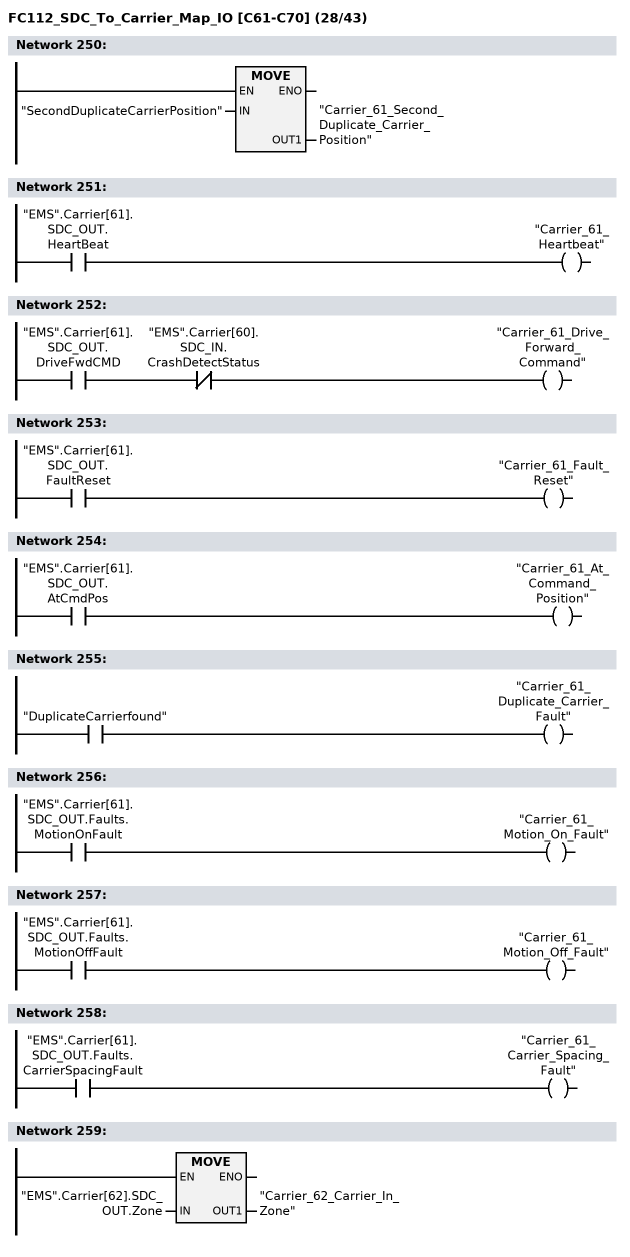
   RUNG wire#powerrail
      Move(in := "SecondDuplicateCarrierPosition", out1 => "Carrier_61_Second_Duplicate_Carrier_Position")
   END_RUNG
   // the same network as SCL:
   "Carrier_61_Second_Duplicate_Carrier_Position" := "SecondDuplicateCarrierPosition";
END_REGION

REGION Network 251
   RUNG wire#powerrail
      Contact( "EMS".Carrier[61].SDC_OUT.HeartBeat )
      Coil( "Carrier_61_Heartbeat" )
   END_RUNG
   // the same network as SCL:
   "Carrier_61_Heartbeat" := "EMS".Carrier[61].SDC_OUT.HeartBeat;
END_REGION

REGION Network 252
   RUNG wire#powerrail
      Contact( "EMS".Carrier[61].SDC_OUT.DriveFwdCMD )
      I_Contact( "EMS".Carrier[60].SDC_IN.CrashDetectStatus )
      Coil( "Carrier_61_Drive_Forward_Command" )
   END_RUNG
   // the same network as SCL:
   "Carrier_61_Drive_Forward_Command" := "EMS".Carrier[61].SDC_OUT.DriveFwdCMD AND NOT "EMS".Carrier[60].SDC_IN.CrashDetectStatus;
END_REGION

REGION Network 253
   RUNG wire#powerrail
      Contact( "EMS".Carrier[61].SDC_OUT.FaultReset )
      Coil( "Carrier_61_Fault_Reset" )
   END_RUNG
   // the same network as SCL:
   "Carrier_61_Fault_Reset" := "EMS".Carrier[61].SDC_OUT.FaultReset;
END_REGION

REGION Network 254
   RUNG wire#powerrail
      Contact( "EMS".Carrier[61].SDC_OUT.AtCmdPos )
      Coil( "Carrier_61_At_Command_Position" )
   END_RUNG
   // the same network as SCL:
   "Carrier_61_At_Command_Position" := "EMS".Carrier[61].SDC_OUT.AtCmdPos;
END_REGION

REGION Network 255
   RUNG wire#powerrail
      Contact( "DuplicateCarrierfound" )
      Coil( "Carrier_61_Duplicate_Carrier_Fault" )
   END_RUNG
   // the same network as SCL:
   "Carrier_61_Duplicate_Carrier_Fault" := "DuplicateCarrierfound";
END_REGION

REGION Network 256
   RUNG wire#powerrail
      Contact( "EMS".Carrier[61].SDC_OUT.Faults.MotionOnFault )
      Coil( "Carrier_61_Motion_On_Fault" )
   END_RUNG
   // the same network as SCL:
   "Carrier_61_Motion_On_Fault" := "EMS".Carrier[61].SDC_OUT.Faults.MotionOnFault;
END_REGION

REGION Network 257
   RUNG wire#powerrail
      Contact( "EMS".Carrier[61].SDC_OUT.Faults.MotionOffFault )
      Coil( "Carrier_61_Motion_Off_Fault" )
   END_RUNG
   // the same network as SCL:
   "Carrier_61_Motion_Off_Fault" := "EMS".Carrier[61].SDC_OUT.Faults.MotionOffFault;
END_REGION

REGION Network 258
   RUNG wire#powerrail
      Contact( "EMS".Carrier[61].SDC_OUT.Faults.CarrierSpacingFault )
      Coil( "Carrier_61_Carrier_Spacing_Fault" )
   END_RUNG
   // the same network as SCL:
   "Carrier_61_Carrier_Spacing_Fault" := "EMS".Carrier[61].SDC_OUT.Faults.CarrierSpacingFault;
END_REGION

REGION Network 259
   RUNG wire#powerrail
      Move(in := "EMS".Carrier[62].SDC_OUT.Zone, out1 => "Carrier_62_Carrier_In_Zone")
   END_RUNG
   // the same network as SCL:
   "Carrier_62_Carrier_In_Zone" := "EMS".Carrier[62].SDC_OUT.Zone;
END_REGION

REGION Network 260
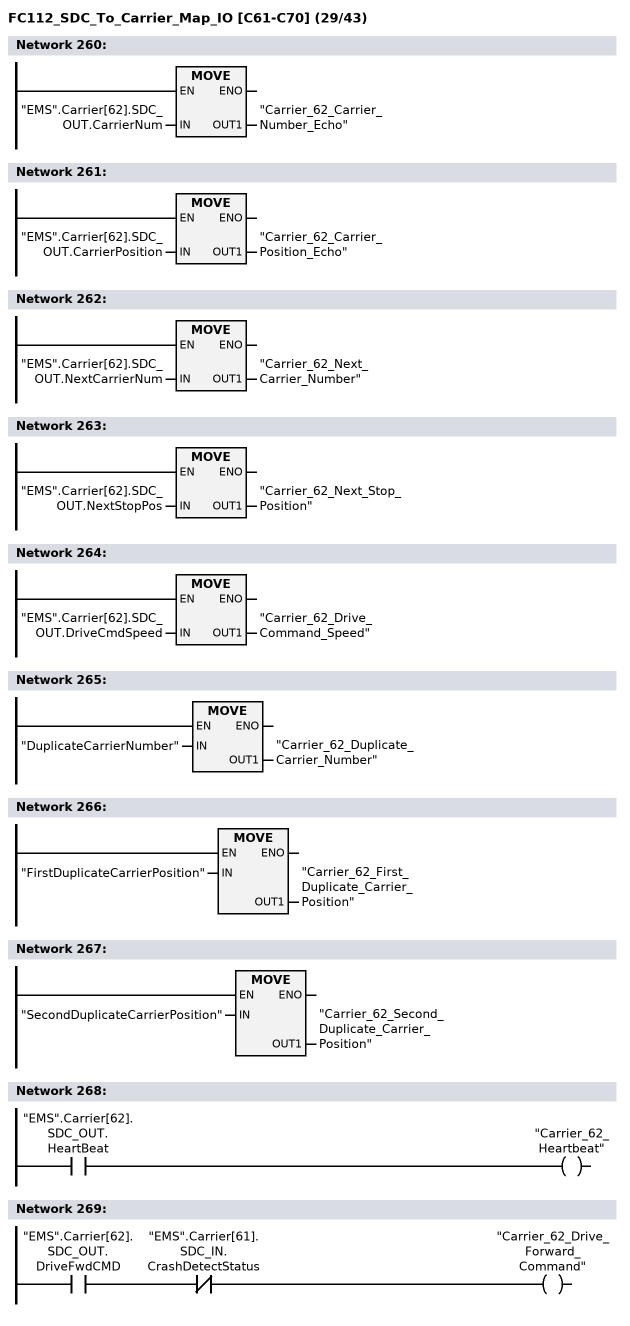
   RUNG wire#powerrail
      Move(in := "EMS".Carrier[62].SDC_OUT.CarrierNum, out1 => "Carrier_62_Carrier_Number_Echo")
   END_RUNG
   // the same network as SCL:
   "Carrier_62_Carrier_Number_Echo" := "EMS".Carrier[62].SDC_OUT.CarrierNum;
END_REGION

REGION Network 261
   RUNG wire#powerrail
      Move(in := "EMS".Carrier[62].SDC_OUT.CarrierPosition, out1 => "Carrier_62_Carrier_Position_Echo")
   END_RUNG
   // the same network as SCL:
   "Carrier_62_Carrier_Position_Echo" := "EMS".Carrier[62].SDC_OUT.CarrierPosition;
END_REGION

REGION Network 262
   RUNG wire#powerrail
      Move(in := "EMS".Carrier[62].SDC_OUT.NextCarrierNum, out1 => "Carrier_62_Next_Carrier_Number")
   END_RUNG
   // the same network as SCL:
   "Carrier_62_Next_Carrier_Number" := "EMS".Carrier[62].SDC_OUT.NextCarrierNum;
END_REGION

REGION Network 263
   RUNG wire#powerrail
      Move(in := "EMS".Carrier[62].SDC_OUT.NextStopPos, out1 => "Carrier_62_Next_Stop_Position")
   END_RUNG
   // the same network as SCL:
   "Carrier_62_Next_Stop_Position" := "EMS".Carrier[62].SDC_OUT.NextStopPos;
END_REGION

REGION Network 264
   RUNG wire#powerrail
      Move(in := "EMS".Carrier[62].SDC_OUT.DriveCmdSpeed, out1 => "Carrier_62_Drive_Command_Speed")
   END_RUNG
   // the same network as SCL:
   "Carrier_62_Drive_Command_Speed" := "EMS".Carrier[62].SDC_OUT.DriveCmdSpeed;
END_REGION

REGION Network 265
   RUNG wire#powerrail
      Move(in := "DuplicateCarrierNumber", out1 => "Carrier_62_Duplicate_Carrier_Number")
   END_RUNG
   // the same network as SCL:
   "Carrier_62_Duplicate_Carrier_Number" := "DuplicateCarrierNumber";
END_REGION

REGION Network 266
   RUNG wire#powerrail
      Move(in := "FirstDuplicateCarrierPosition", out1 => "Carrier_62_First_Duplicate_Carrier_Position")
   END_RUNG
   // the same network as SCL:
   "Carrier_62_First_Duplicate_Carrier_Position" := "FirstDuplicateCarrierPosition";
END_REGION

REGION Network 267
   RUNG wire#powerrail
      Move(in := "SecondDuplicateCarrierPosition", out1 => "Carrier_62_Second_Duplicate_Carrier_Position")
   END_RUNG
   // the same network as SCL:
   "Carrier_62_Second_Duplicate_Carrier_Position" := "SecondDuplicateCarrierPosition";
END_REGION

REGION Network 268
   RUNG wire#powerrail
      Contact( "EMS".Carrier[62].SDC_OUT.HeartBeat )
      Coil( "Carrier_62_Heartbeat" )
   END_RUNG
   // the same network as SCL:
   "Carrier_62_Heartbeat" := "EMS".Carrier[62].SDC_OUT.HeartBeat;
END_REGION

REGION Network 269
   RUNG wire#powerrail
      Contact( "EMS".Carrier[62].SDC_OUT.DriveFwdCMD )
      I_Contact( "EMS".Carrier[61].SDC_IN.CrashDetectStatus )
      Coil( "Carrier_62_Drive_Forward_Command" )
   END_RUNG
   // the same network as SCL:
   "Carrier_62_Drive_Forward_Command" := "EMS".Carrier[62].SDC_OUT.DriveFwdCMD AND NOT "EMS".Carrier[61].SDC_IN.CrashDetectStatus;
END_REGION

REGION Network 270
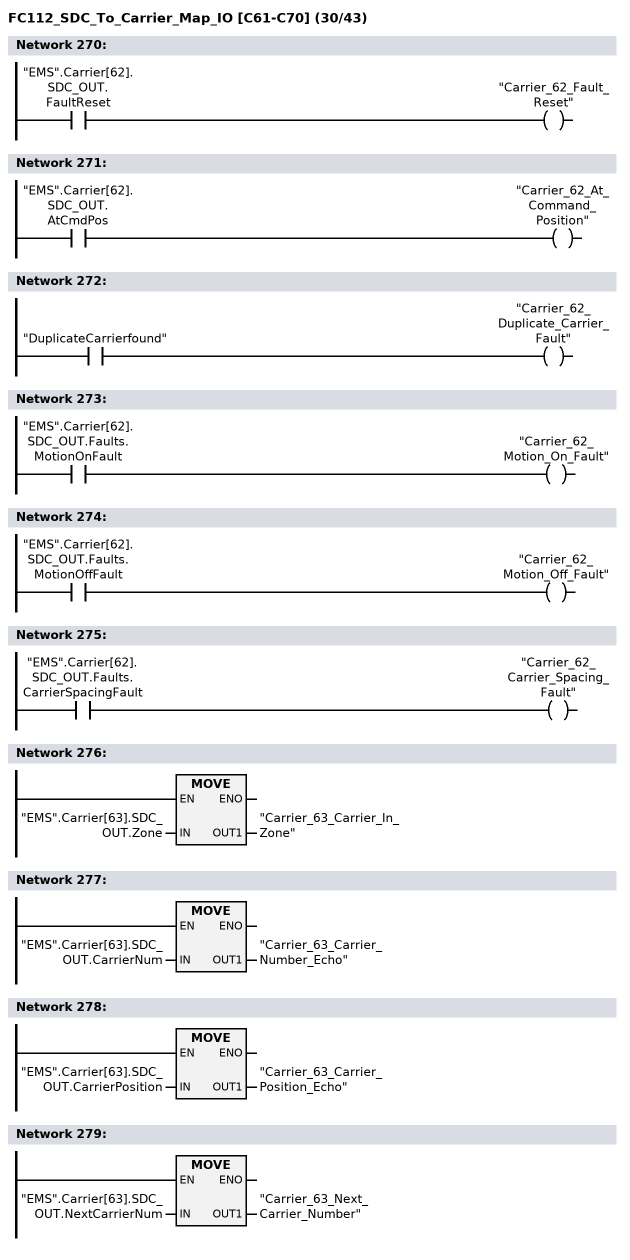
   RUNG wire#powerrail
      Contact( "EMS".Carrier[62].SDC_OUT.FaultReset )
      Coil( "Carrier_62_Fault_Reset" )
   END_RUNG
   // the same network as SCL:
   "Carrier_62_Fault_Reset" := "EMS".Carrier[62].SDC_OUT.FaultReset;
END_REGION

REGION Network 271
   RUNG wire#powerrail
      Contact( "EMS".Carrier[62].SDC_OUT.AtCmdPos )
      Coil( "Carrier_62_At_Command_Position" )
   END_RUNG
   // the same network as SCL:
   "Carrier_62_At_Command_Position" := "EMS".Carrier[62].SDC_OUT.AtCmdPos;
END_REGION

REGION Network 272
   RUNG wire#powerrail
      Contact( "DuplicateCarrierfound" )
      Coil( "Carrier_62_Duplicate_Carrier_Fault" )
   END_RUNG
   // the same network as SCL:
   "Carrier_62_Duplicate_Carrier_Fault" := "DuplicateCarrierfound";
END_REGION

REGION Network 273
   RUNG wire#powerrail
      Contact( "EMS".Carrier[62].SDC_OUT.Faults.MotionOnFault )
      Coil( "Carrier_62_Motion_On_Fault" )
   END_RUNG
   // the same network as SCL:
   "Carrier_62_Motion_On_Fault" := "EMS".Carrier[62].SDC_OUT.Faults.MotionOnFault;
END_REGION

REGION Network 274
   RUNG wire#powerrail
      Contact( "EMS".Carrier[62].SDC_OUT.Faults.MotionOffFault )
      Coil( "Carrier_62_Motion_Off_Fault" )
   END_RUNG
   // the same network as SCL:
   "Carrier_62_Motion_Off_Fault" := "EMS".Carrier[62].SDC_OUT.Faults.MotionOffFault;
END_REGION

REGION Network 275
   RUNG wire#powerrail
      Contact( "EMS".Carrier[62].SDC_OUT.Faults.CarrierSpacingFault )
      Coil( "Carrier_62_Carrier_Spacing_Fault" )
   END_RUNG
   // the same network as SCL:
   "Carrier_62_Carrier_Spacing_Fault" := "EMS".Carrier[62].SDC_OUT.Faults.CarrierSpacingFault;
END_REGION

REGION Network 276
   RUNG wire#powerrail
      Move(in := "EMS".Carrier[63].SDC_OUT.Zone, out1 => "Carrier_63_Carrier_In_Zone")
   END_RUNG
   // the same network as SCL:
   "Carrier_63_Carrier_In_Zone" := "EMS".Carrier[63].SDC_OUT.Zone;
END_REGION

REGION Network 277
   RUNG wire#powerrail
      Move(in := "EMS".Carrier[63].SDC_OUT.CarrierNum, out1 => "Carrier_63_Carrier_Number_Echo")
   END_RUNG
   // the same network as SCL:
   "Carrier_63_Carrier_Number_Echo" := "EMS".Carrier[63].SDC_OUT.CarrierNum;
END_REGION

REGION Network 278
   RUNG wire#powerrail
      Move(in := "EMS".Carrier[63].SDC_OUT.CarrierPosition, out1 => "Carrier_63_Carrier_Position_Echo")
   END_RUNG
   // the same network as SCL:
   "Carrier_63_Carrier_Position_Echo" := "EMS".Carrier[63].SDC_OUT.CarrierPosition;
END_REGION

REGION Network 279
   RUNG wire#powerrail
      Move(in := "EMS".Carrier[63].SDC_OUT.NextCarrierNum, out1 => "Carrier_63_Next_Carrier_Number")
   END_RUNG
   // the same network as SCL:
   "Carrier_63_Next_Carrier_Number" := "EMS".Carrier[63].SDC_OUT.NextCarrierNum;
END_REGION

REGION Network 280
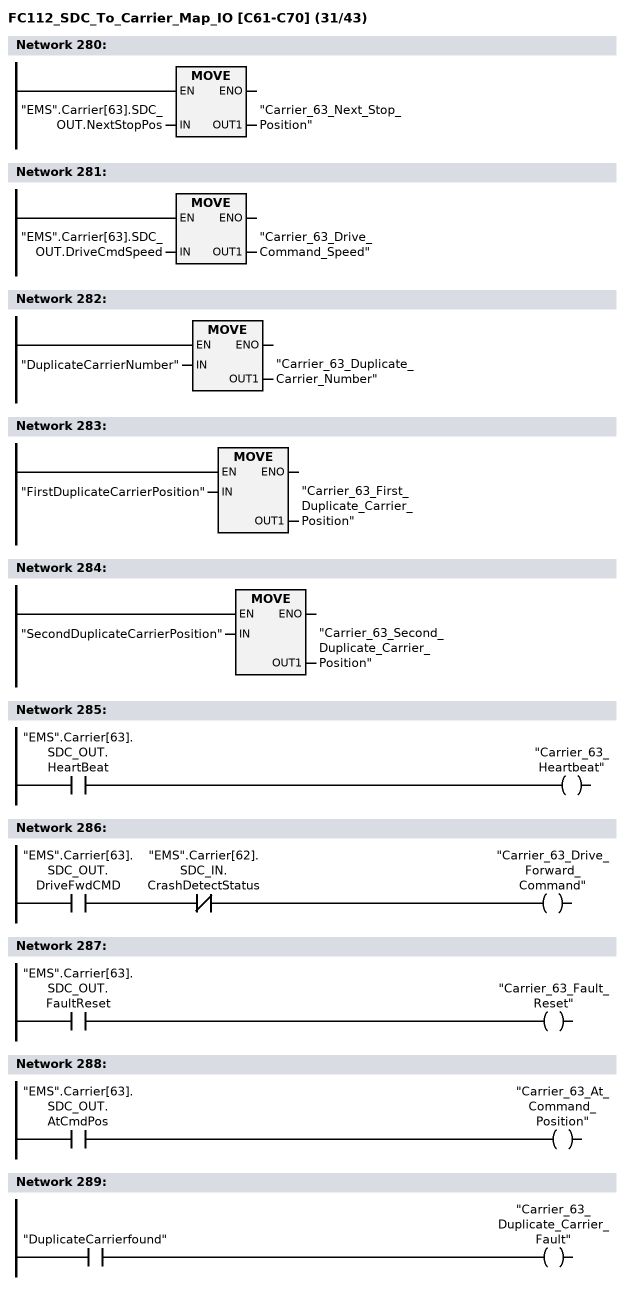
   RUNG wire#powerrail
      Move(in := "EMS".Carrier[63].SDC_OUT.NextStopPos, out1 => "Carrier_63_Next_Stop_Position")
   END_RUNG
   // the same network as SCL:
   "Carrier_63_Next_Stop_Position" := "EMS".Carrier[63].SDC_OUT.NextStopPos;
END_REGION

REGION Network 281
   RUNG wire#powerrail
      Move(in := "EMS".Carrier[63].SDC_OUT.DriveCmdSpeed, out1 => "Carrier_63_Drive_Command_Speed")
   END_RUNG
   // the same network as SCL:
   "Carrier_63_Drive_Command_Speed" := "EMS".Carrier[63].SDC_OUT.DriveCmdSpeed;
END_REGION

REGION Network 282
   RUNG wire#powerrail
      Move(in := "DuplicateCarrierNumber", out1 => "Carrier_63_Duplicate_Carrier_Number")
   END_RUNG
   // the same network as SCL:
   "Carrier_63_Duplicate_Carrier_Number" := "DuplicateCarrierNumber";
END_REGION

REGION Network 283
   RUNG wire#powerrail
      Move(in := "FirstDuplicateCarrierPosition", out1 => "Carrier_63_First_Duplicate_Carrier_Position")
   END_RUNG
   // the same network as SCL:
   "Carrier_63_First_Duplicate_Carrier_Position" := "FirstDuplicateCarrierPosition";
END_REGION

REGION Network 284
   RUNG wire#powerrail
      Move(in := "SecondDuplicateCarrierPosition", out1 => "Carrier_63_Second_Duplicate_Carrier_Position")
   END_RUNG
   // the same network as SCL:
   "Carrier_63_Second_Duplicate_Carrier_Position" := "SecondDuplicateCarrierPosition";
END_REGION

REGION Network 285
   RUNG wire#powerrail
      Contact( "EMS".Carrier[63].SDC_OUT.HeartBeat )
      Coil( "Carrier_63_Heartbeat" )
   END_RUNG
   // the same network as SCL:
   "Carrier_63_Heartbeat" := "EMS".Carrier[63].SDC_OUT.HeartBeat;
END_REGION

REGION Network 286
   RUNG wire#powerrail
      Contact( "EMS".Carrier[63].SDC_OUT.DriveFwdCMD )
      I_Contact( "EMS".Carrier[62].SDC_IN.CrashDetectStatus )
      Coil( "Carrier_63_Drive_Forward_Command" )
   END_RUNG
   // the same network as SCL:
   "Carrier_63_Drive_Forward_Command" := "EMS".Carrier[63].SDC_OUT.DriveFwdCMD AND NOT "EMS".Carrier[62].SDC_IN.CrashDetectStatus;
END_REGION

REGION Network 287
   RUNG wire#powerrail
      Contact( "EMS".Carrier[63].SDC_OUT.FaultReset )
      Coil( "Carrier_63_Fault_Reset" )
   END_RUNG
   // the same network as SCL:
   "Carrier_63_Fault_Reset" := "EMS".Carrier[63].SDC_OUT.FaultReset;
END_REGION

REGION Network 288
   RUNG wire#powerrail
      Contact( "EMS".Carrier[63].SDC_OUT.AtCmdPos )
      Coil( "Carrier_63_At_Command_Position" )
   END_RUNG
   // the same network as SCL:
   "Carrier_63_At_Command_Position" := "EMS".Carrier[63].SDC_OUT.AtCmdPos;
END_REGION

REGION Network 289
   RUNG wire#powerrail
      Contact( "DuplicateCarrierfound" )
      Coil( "Carrier_63_Duplicate_Carrier_Fault" )
   END_RUNG
   // the same network as SCL:
   "Carrier_63_Duplicate_Carrier_Fault" := "DuplicateCarrierfound";
END_REGION

REGION Network 290
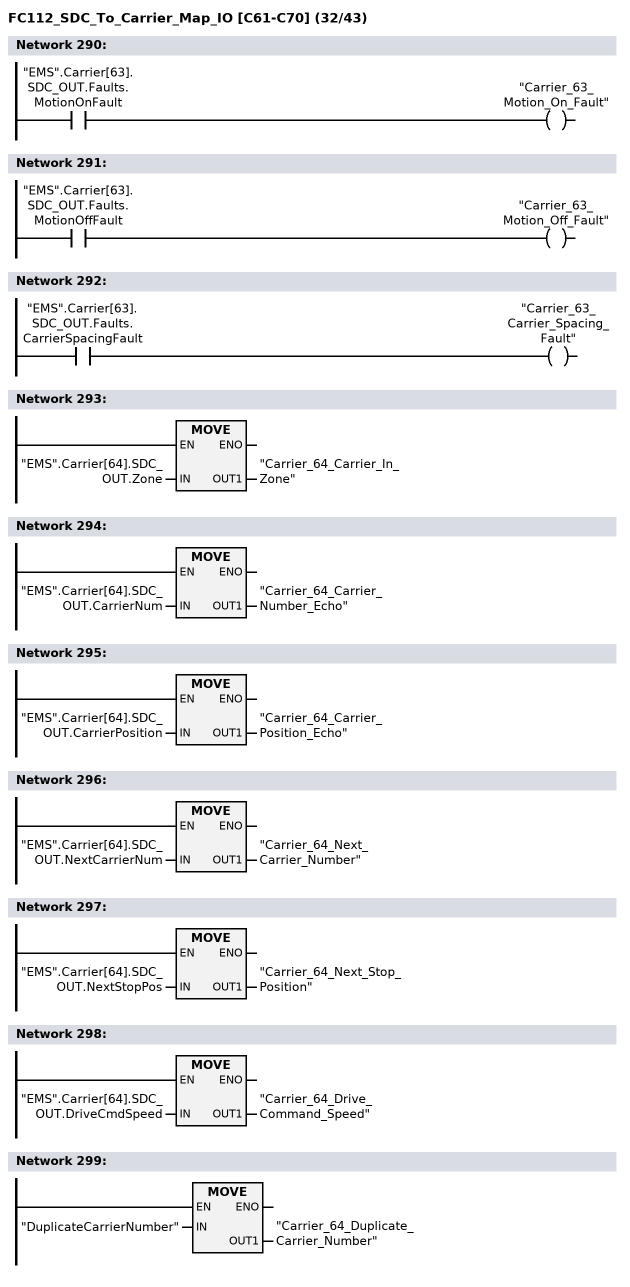
   RUNG wire#powerrail
      Contact( "EMS".Carrier[63].SDC_OUT.Faults.MotionOnFault )
      Coil( "Carrier_63_Motion_On_Fault" )
   END_RUNG
   // the same network as SCL:
   "Carrier_63_Motion_On_Fault" := "EMS".Carrier[63].SDC_OUT.Faults.MotionOnFault;
END_REGION

REGION Network 291
   RUNG wire#powerrail
      Contact( "EMS".Carrier[63].SDC_OUT.Faults.MotionOffFault )
      Coil( "Carrier_63_Motion_Off_Fault" )
   END_RUNG
   // the same network as SCL:
   "Carrier_63_Motion_Off_Fault" := "EMS".Carrier[63].SDC_OUT.Faults.MotionOffFault;
END_REGION

REGION Network 292
   RUNG wire#powerrail
      Contact( "EMS".Carrier[63].SDC_OUT.Faults.CarrierSpacingFault )
      Coil( "Carrier_63_Carrier_Spacing_Fault" )
   END_RUNG
   // the same network as SCL:
   "Carrier_63_Carrier_Spacing_Fault" := "EMS".Carrier[63].SDC_OUT.Faults.CarrierSpacingFault;
END_REGION

REGION Network 293
   RUNG wire#powerrail
      Move(in := "EMS".Carrier[64].SDC_OUT.Zone, out1 => "Carrier_64_Carrier_In_Zone")
   END_RUNG
   // the same network as SCL:
   "Carrier_64_Carrier_In_Zone" := "EMS".Carrier[64].SDC_OUT.Zone;
END_REGION

REGION Network 294
   RUNG wire#powerrail
      Move(in := "EMS".Carrier[64].SDC_OUT.CarrierNum, out1 => "Carrier_64_Carrier_Number_Echo")
   END_RUNG
   // the same network as SCL:
   "Carrier_64_Carrier_Number_Echo" := "EMS".Carrier[64].SDC_OUT.CarrierNum;
END_REGION

REGION Network 295
   RUNG wire#powerrail
      Move(in := "EMS".Carrier[64].SDC_OUT.CarrierPosition, out1 => "Carrier_64_Carrier_Position_Echo")
   END_RUNG
   // the same network as SCL:
   "Carrier_64_Carrier_Position_Echo" := "EMS".Carrier[64].SDC_OUT.CarrierPosition;
END_REGION

REGION Network 296
   RUNG wire#powerrail
      Move(in := "EMS".Carrier[64].SDC_OUT.NextCarrierNum, out1 => "Carrier_64_Next_Carrier_Number")
   END_RUNG
   // the same network as SCL:
   "Carrier_64_Next_Carrier_Number" := "EMS".Carrier[64].SDC_OUT.NextCarrierNum;
END_REGION

REGION Network 297
   RUNG wire#powerrail
      Move(in := "EMS".Carrier[64].SDC_OUT.NextStopPos, out1 => "Carrier_64_Next_Stop_Position")
   END_RUNG
   // the same network as SCL:
   "Carrier_64_Next_Stop_Position" := "EMS".Carrier[64].SDC_OUT.NextStopPos;
END_REGION

REGION Network 298
   RUNG wire#powerrail
      Move(in := "EMS".Carrier[64].SDC_OUT.DriveCmdSpeed, out1 => "Carrier_64_Drive_Command_Speed")
   END_RUNG
   // the same network as SCL:
   "Carrier_64_Drive_Command_Speed" := "EMS".Carrier[64].SDC_OUT.DriveCmdSpeed;
END_REGION

REGION Network 299
   RUNG wire#powerrail
      Move(in := "DuplicateCarrierNumber", out1 => "Carrier_64_Duplicate_Carrier_Number")
   END_RUNG
   // the same network as SCL:
   "Carrier_64_Duplicate_Carrier_Number" := "DuplicateCarrierNumber";
END_REGION

REGION Network 300
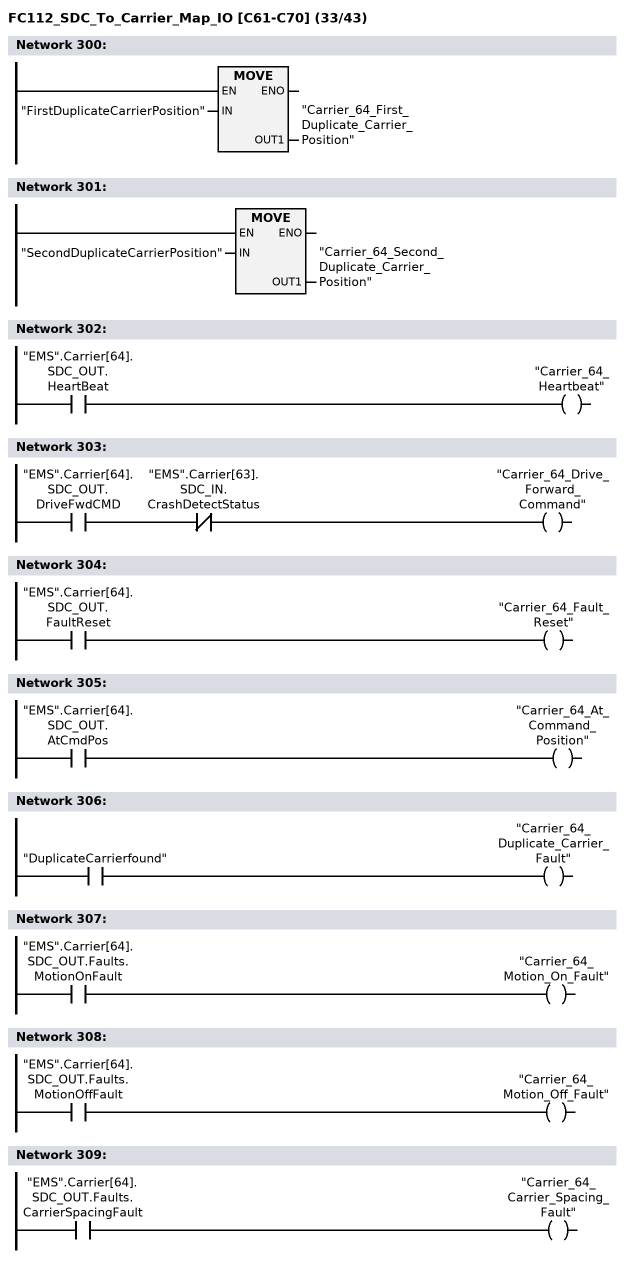
   RUNG wire#powerrail
      Move(in := "FirstDuplicateCarrierPosition", out1 => "Carrier_64_First_Duplicate_Carrier_Position")
   END_RUNG
   // the same network as SCL:
   "Carrier_64_First_Duplicate_Carrier_Position" := "FirstDuplicateCarrierPosition";
END_REGION

REGION Network 301
   RUNG wire#powerrail
      Move(in := "SecondDuplicateCarrierPosition", out1 => "Carrier_64_Second_Duplicate_Carrier_Position")
   END_RUNG
   // the same network as SCL:
   "Carrier_64_Second_Duplicate_Carrier_Position" := "SecondDuplicateCarrierPosition";
END_REGION

REGION Network 302
   RUNG wire#powerrail
      Contact( "EMS".Carrier[64].SDC_OUT.HeartBeat )
      Coil( "Carrier_64_Heartbeat" )
   END_RUNG
   // the same network as SCL:
   "Carrier_64_Heartbeat" := "EMS".Carrier[64].SDC_OUT.HeartBeat;
END_REGION

REGION Network 303
   RUNG wire#powerrail
      Contact( "EMS".Carrier[64].SDC_OUT.DriveFwdCMD )
      I_Contact( "EMS".Carrier[63].SDC_IN.CrashDetectStatus )
      Coil( "Carrier_64_Drive_Forward_Command" )
   END_RUNG
   // the same network as SCL:
   "Carrier_64_Drive_Forward_Command" := "EMS".Carrier[64].SDC_OUT.DriveFwdCMD AND NOT "EMS".Carrier[63].SDC_IN.CrashDetectStatus;
END_REGION

REGION Network 304
   RUNG wire#powerrail
      Contact( "EMS".Carrier[64].SDC_OUT.FaultReset )
      Coil( "Carrier_64_Fault_Reset" )
   END_RUNG
   // the same network as SCL:
   "Carrier_64_Fault_Reset" := "EMS".Carrier[64].SDC_OUT.FaultReset;
END_REGION

REGION Network 305
   RUNG wire#powerrail
      Contact( "EMS".Carrier[64].SDC_OUT.AtCmdPos )
      Coil( "Carrier_64_At_Command_Position" )
   END_RUNG
   // the same network as SCL:
   "Carrier_64_At_Command_Position" := "EMS".Carrier[64].SDC_OUT.AtCmdPos;
END_REGION

REGION Network 306
   RUNG wire#powerrail
      Contact( "DuplicateCarrierfound" )
      Coil( "Carrier_64_Duplicate_Carrier_Fault" )
   END_RUNG
   // the same network as SCL:
   "Carrier_64_Duplicate_Carrier_Fault" := "DuplicateCarrierfound";
END_REGION

REGION Network 307
   RUNG wire#powerrail
      Contact( "EMS".Carrier[64].SDC_OUT.Faults.MotionOnFault )
      Coil( "Carrier_64_Motion_On_Fault" )
   END_RUNG
   // the same network as SCL:
   "Carrier_64_Motion_On_Fault" := "EMS".Carrier[64].SDC_OUT.Faults.MotionOnFault;
END_REGION

REGION Network 308
   RUNG wire#powerrail
      Contact( "EMS".Carrier[64].SDC_OUT.Faults.MotionOffFault )
      Coil( "Carrier_64_Motion_Off_Fault" )
   END_RUNG
   // the same network as SCL:
   "Carrier_64_Motion_Off_Fault" := "EMS".Carrier[64].SDC_OUT.Faults.MotionOffFault;
END_REGION

REGION Network 309
   RUNG wire#powerrail
      Contact( "EMS".Carrier[64].SDC_OUT.Faults.CarrierSpacingFault )
      Coil( "Carrier_64_Carrier_Spacing_Fault" )
   END_RUNG
   // the same network as SCL:
   "Carrier_64_Carrier_Spacing_Fault" := "EMS".Carrier[64].SDC_OUT.Faults.CarrierSpacingFault;
END_REGION

REGION Network 310
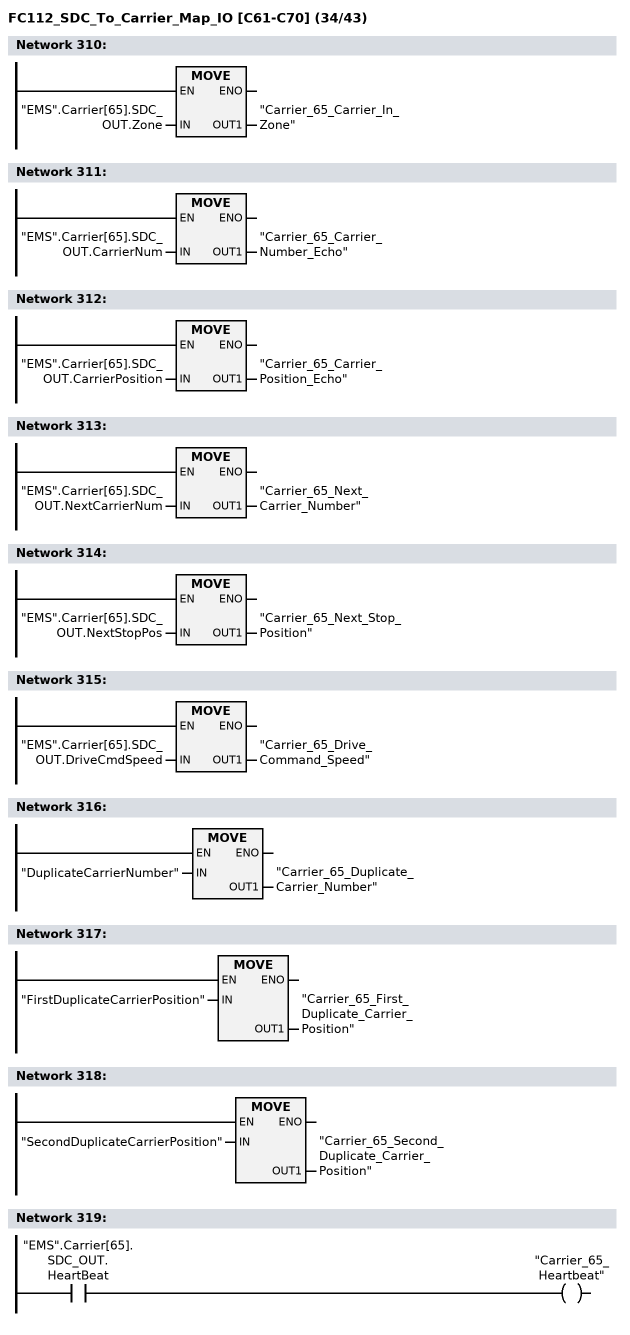
   RUNG wire#powerrail
      Move(in := "EMS".Carrier[65].SDC_OUT.Zone, out1 => "Carrier_65_Carrier_In_Zone")
   END_RUNG
   // the same network as SCL:
   "Carrier_65_Carrier_In_Zone" := "EMS".Carrier[65].SDC_OUT.Zone;
END_REGION

REGION Network 311
   RUNG wire#powerrail
      Move(in := "EMS".Carrier[65].SDC_OUT.CarrierNum, out1 => "Carrier_65_Carrier_Number_Echo")
   END_RUNG
   // the same network as SCL:
   "Carrier_65_Carrier_Number_Echo" := "EMS".Carrier[65].SDC_OUT.CarrierNum;
END_REGION

REGION Network 312
   RUNG wire#powerrail
      Move(in := "EMS".Carrier[65].SDC_OUT.CarrierPosition, out1 => "Carrier_65_Carrier_Position_Echo")
   END_RUNG
   // the same network as SCL:
   "Carrier_65_Carrier_Position_Echo" := "EMS".Carrier[65].SDC_OUT.CarrierPosition;
END_REGION

REGION Network 313
   RUNG wire#powerrail
      Move(in := "EMS".Carrier[65].SDC_OUT.NextCarrierNum, out1 => "Carrier_65_Next_Carrier_Number")
   END_RUNG
   // the same network as SCL:
   "Carrier_65_Next_Carrier_Number" := "EMS".Carrier[65].SDC_OUT.NextCarrierNum;
END_REGION

REGION Network 314
   RUNG wire#powerrail
      Move(in := "EMS".Carrier[65].SDC_OUT.NextStopPos, out1 => "Carrier_65_Next_Stop_Position")
   END_RUNG
   // the same network as SCL:
   "Carrier_65_Next_Stop_Position" := "EMS".Carrier[65].SDC_OUT.NextStopPos;
END_REGION

REGION Network 315
   RUNG wire#powerrail
      Move(in := "EMS".Carrier[65].SDC_OUT.DriveCmdSpeed, out1 => "Carrier_65_Drive_Command_Speed")
   END_RUNG
   // the same network as SCL:
   "Carrier_65_Drive_Command_Speed" := "EMS".Carrier[65].SDC_OUT.DriveCmdSpeed;
END_REGION

REGION Network 316
   RUNG wire#powerrail
      Move(in := "DuplicateCarrierNumber", out1 => "Carrier_65_Duplicate_Carrier_Number")
   END_RUNG
   // the same network as SCL:
   "Carrier_65_Duplicate_Carrier_Number" := "DuplicateCarrierNumber";
END_REGION

REGION Network 317
   RUNG wire#powerrail
      Move(in := "FirstDuplicateCarrierPosition", out1 => "Carrier_65_First_Duplicate_Carrier_Position")
   END_RUNG
   // the same network as SCL:
   "Carrier_65_First_Duplicate_Carrier_Position" := "FirstDuplicateCarrierPosition";
END_REGION

REGION Network 318
   RUNG wire#powerrail
      Move(in := "SecondDuplicateCarrierPosition", out1 => "Carrier_65_Second_Duplicate_Carrier_Position")
   END_RUNG
   // the same network as SCL:
   "Carrier_65_Second_Duplicate_Carrier_Position" := "SecondDuplicateCarrierPosition";
END_REGION

REGION Network 319
   RUNG wire#powerrail
      Contact( "EMS".Carrier[65].SDC_OUT.HeartBeat )
      Coil( "Carrier_65_Heartbeat" )
   END_RUNG
   // the same network as SCL:
   "Carrier_65_Heartbeat" := "EMS".Carrier[65].SDC_OUT.HeartBeat;
END_REGION

REGION Network 320
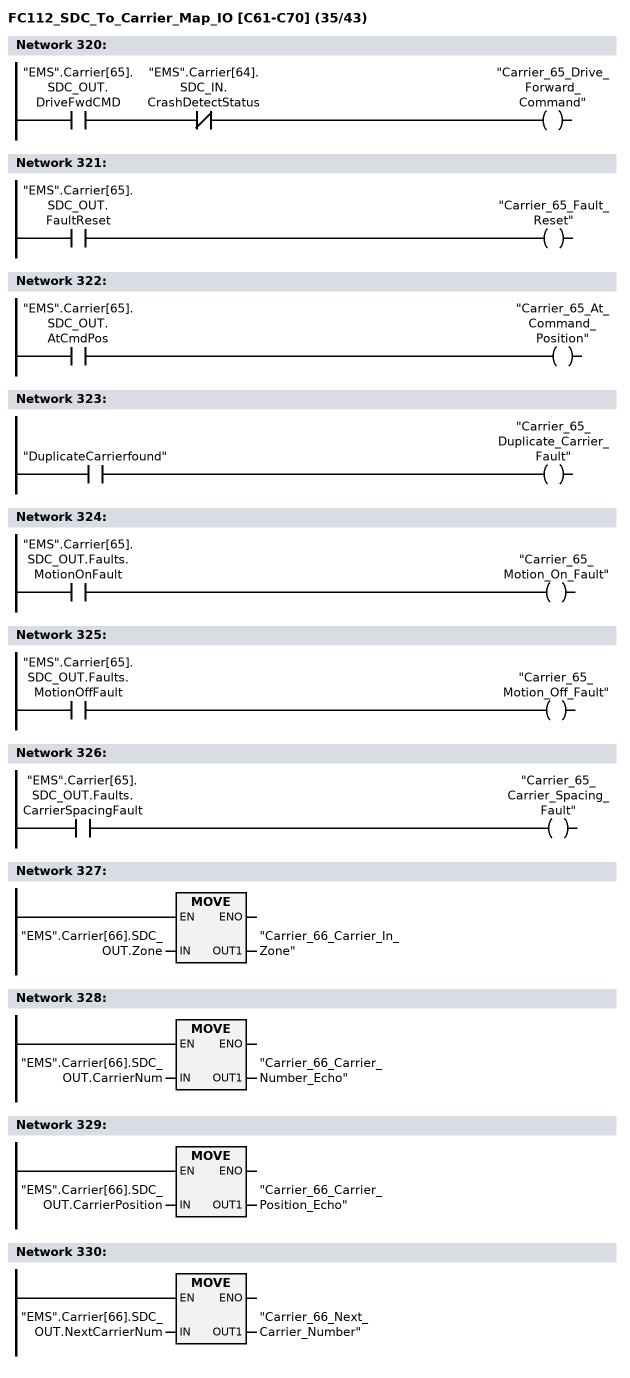
   RUNG wire#powerrail
      Contact( "EMS".Carrier[65].SDC_OUT.DriveFwdCMD )
      I_Contact( "EMS".Carrier[64].SDC_IN.CrashDetectStatus )
      Coil( "Carrier_65_Drive_Forward_Command" )
   END_RUNG
   // the same network as SCL:
   "Carrier_65_Drive_Forward_Command" := "EMS".Carrier[65].SDC_OUT.DriveFwdCMD AND NOT "EMS".Carrier[64].SDC_IN.CrashDetectStatus;
END_REGION

REGION Network 321
   RUNG wire#powerrail
      Contact( "EMS".Carrier[65].SDC_OUT.FaultReset )
      Coil( "Carrier_65_Fault_Reset" )
   END_RUNG
   // the same network as SCL:
   "Carrier_65_Fault_Reset" := "EMS".Carrier[65].SDC_OUT.FaultReset;
END_REGION

REGION Network 322
   RUNG wire#powerrail
      Contact( "EMS".Carrier[65].SDC_OUT.AtCmdPos )
      Coil( "Carrier_65_At_Command_Position" )
   END_RUNG
   // the same network as SCL:
   "Carrier_65_At_Command_Position" := "EMS".Carrier[65].SDC_OUT.AtCmdPos;
END_REGION

REGION Network 323
   RUNG wire#powerrail
      Contact( "DuplicateCarrierfound" )
      Coil( "Carrier_65_Duplicate_Carrier_Fault" )
   END_RUNG
   // the same network as SCL:
   "Carrier_65_Duplicate_Carrier_Fault" := "DuplicateCarrierfound";
END_REGION

REGION Network 324
   RUNG wire#powerrail
      Contact( "EMS".Carrier[65].SDC_OUT.Faults.MotionOnFault )
      Coil( "Carrier_65_Motion_On_Fault" )
   END_RUNG
   // the same network as SCL:
   "Carrier_65_Motion_On_Fault" := "EMS".Carrier[65].SDC_OUT.Faults.MotionOnFault;
END_REGION

REGION Network 325
   RUNG wire#powerrail
      Contact( "EMS".Carrier[65].SDC_OUT.Faults.MotionOffFault )
      Coil( "Carrier_65_Motion_Off_Fault" )
   END_RUNG
   // the same network as SCL:
   "Carrier_65_Motion_Off_Fault" := "EMS".Carrier[65].SDC_OUT.Faults.MotionOffFault;
END_REGION

REGION Network 326
   RUNG wire#powerrail
      Contact( "EMS".Carrier[65].SDC_OUT.Faults.CarrierSpacingFault )
      Coil( "Carrier_65_Carrier_Spacing_Fault" )
   END_RUNG
   // the same network as SCL:
   "Carrier_65_Carrier_Spacing_Fault" := "EMS".Carrier[65].SDC_OUT.Faults.CarrierSpacingFault;
END_REGION

REGION Network 327
   RUNG wire#powerrail
      Move(in := "EMS".Carrier[66].SDC_OUT.Zone, out1 => "Carrier_66_Carrier_In_Zone")
   END_RUNG
   // the same network as SCL:
   "Carrier_66_Carrier_In_Zone" := "EMS".Carrier[66].SDC_OUT.Zone;
END_REGION

REGION Network 328
   RUNG wire#powerrail
      Move(in := "EMS".Carrier[66].SDC_OUT.CarrierNum, out1 => "Carrier_66_Carrier_Number_Echo")
   END_RUNG
   // the same network as SCL:
   "Carrier_66_Carrier_Number_Echo" := "EMS".Carrier[66].SDC_OUT.CarrierNum;
END_REGION

REGION Network 329
   RUNG wire#powerrail
      Move(in := "EMS".Carrier[66].SDC_OUT.CarrierPosition, out1 => "Carrier_66_Carrier_Position_Echo")
   END_RUNG
   // the same network as SCL:
   "Carrier_66_Carrier_Position_Echo" := "EMS".Carrier[66].SDC_OUT.CarrierPosition;
END_REGION

REGION Network 330
   RUNG wire#powerrail
      Move(in := "EMS".Carrier[66].SDC_OUT.NextCarrierNum, out1 => "Carrier_66_Next_Carrier_Number")
   END_RUNG
   // the same network as SCL:
   "Carrier_66_Next_Carrier_Number" := "EMS".Carrier[66].SDC_OUT.NextCarrierNum;
END_REGION

REGION Network 331
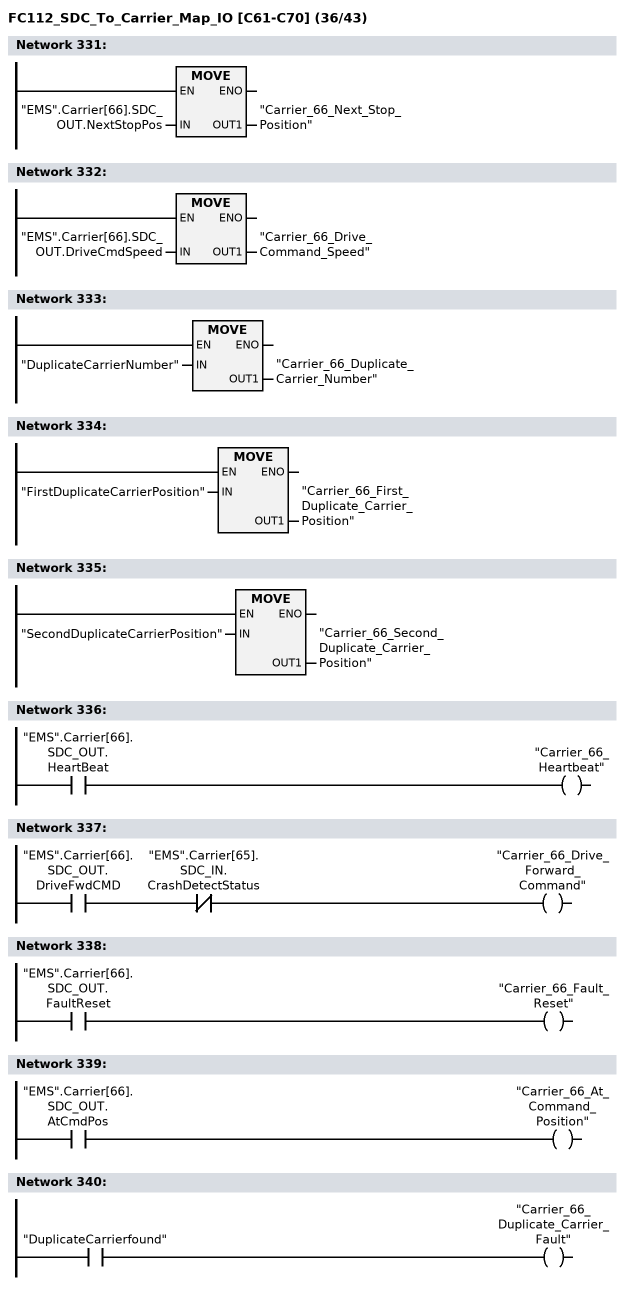
   RUNG wire#powerrail
      Move(in := "EMS".Carrier[66].SDC_OUT.NextStopPos, out1 => "Carrier_66_Next_Stop_Position")
   END_RUNG
   // the same network as SCL:
   "Carrier_66_Next_Stop_Position" := "EMS".Carrier[66].SDC_OUT.NextStopPos;
END_REGION

REGION Network 332
   RUNG wire#powerrail
      Move(in := "EMS".Carrier[66].SDC_OUT.DriveCmdSpeed, out1 => "Carrier_66_Drive_Command_Speed")
   END_RUNG
   // the same network as SCL:
   "Carrier_66_Drive_Command_Speed" := "EMS".Carrier[66].SDC_OUT.DriveCmdSpeed;
END_REGION
